(* Logix 5000 project; controller UOWHF_Vary Emulate 5570 rev 30.12; software revision 30.00; part 2 of 13 *)
(* tags used below, declared in another part *)
   UOWHF_Add_c : DINT;
   UOWHF_Msg : DINT[16];
   UOWHF_OutputMaxInd : DINT;
   UOWHF_Result : DINT[17];
(* MainProgram, continued *)

   		UOWHF_Result[2]:=UOWHF_Result[2] + 2135853958+UOWHF_Add_c;
   		UOWHF_Add_c.2:=UOWHF_Result[2].31;
   		UOWHF_Result[2].31:=0;
   		UOWHF_Result[3]:=UOWHF_Result[3] + 1732375759+UOWHF_Add_c;
   		UOWHF_Add_c.3:=UOWHF_Result[3].31;
   		UOWHF_Result[3].31:=0;
   		UOWHF_Result[4]:=UOWHF_Result[4] + 115158473+UOWHF_Add_c;
   		UOWHF_Add_c.4:=UOWHF_Result[4].31;
   		UOWHF_Result[4].31:=0;
   	End_If;
   	If UOWHF_Msg[4].[8] Then
   		UOWHF_Result[0]:=UOWHF_Result[0] + 1989798588+UOWHF_Add_c;
   		UOWHF_Add_c.0:=UOWHF_Result[0].31;
   		UOWHF_Result[0].31:=0;
   		UOWHF_Result[1]:=UOWHF_Result[1] + 591703516+UOWHF_Add_c;
   		UOWHF_Add_c.1:=UOWHF_Result[1].31;
   		UOWHF_Result[1].31:=0;
   		UOWHF_Result[2]:=UOWHF_Result[2] + 1328366246+UOWHF_Add_c;
   		UOWHF_Add_c.2:=UOWHF_Result[2].31;
   		UOWHF_Result[2].31:=0;
   		UOWHF_Result[3]:=UOWHF_Result[3] + 1055479196+UOWHF_Add_c;
   		UOWHF_Add_c.3:=UOWHF_Result[3].31;
   		UOWHF_Result[3].31:=0;
   		UOWHF_Result[4]:=UOWHF_Result[4] + 1638831242+UOWHF_Add_c;
   		UOWHF_Add_c.4:=UOWHF_Result[4].31;
   		UOWHF_Result[4].31:=0;
   	End_If;
   	If UOWHF_Msg[4].[9] Then
   		UOWHF_Result[0]:=UOWHF_Result[0] + 622406376+UOWHF_Add_c;
   		UOWHF_Add_c.0:=UOWHF_Result[0].31;
   		UOWHF_Result[0].31:=0;
   		UOWHF_Result[1]:=UOWHF_Result[1] + 302456745+UOWHF_Add_c;
   		UOWHF_Add_c.1:=UOWHF_Result[1].31;
   		UOWHF_Result[1].31:=0;
   		UOWHF_Result[2]:=UOWHF_Result[2] + 1004502914+UOWHF_Add_c;
   		UOWHF_Add_c.2:=UOWHF_Result[2].31;
   		UOWHF_Result[2].31:=0;
   		UOWHF_Result[3]:=UOWHF_Result[3] + 1944958998+UOWHF_Add_c;
   		UOWHF_Add_c.3:=UOWHF_Result[3].31;
   		UOWHF_Result[3].31:=0;
   		UOWHF_Result[4]:=UOWHF_Result[4] + 1457990763+UOWHF_Add_c;
   		UOWHF_Add_c.4:=UOWHF_Result[4].31;
   		UOWHF_Result[4].31:=0;
   	End_If;
   	If UOWHF_Msg[4].[10] Then
   		UOWHF_Result[0]:=UOWHF_Result[0] + 1190952435+UOWHF_Add_c;
   		UOWHF_Add_c.0:=UOWHF_Result[0].31;
   		UOWHF_Result[0].31:=0;
   		UOWHF_Result[1]:=UOWHF_Result[1] + 906321176+UOWHF_Add_c;
   		UOWHF_Add_c.1:=UOWHF_Result[1].31;
   		UOWHF_Result[1].31:=0;
   		UOWHF_Result[2]:=UOWHF_Result[2] + 1114856499+UOWHF_Add_c;
   		UOWHF_Add_c.2:=UOWHF_Result[2].31;
   		UOWHF_Result[2].31:=0;
   		UOWHF_Result[3]:=UOWHF_Result[3] + 2109990137+UOWHF_Add_c;
   		UOWHF_Add_c.3:=UOWHF_Result[3].31;
   		UOWHF_Result[3].31:=0;
   		UOWHF_Result[4]:=UOWHF_Result[4] + 2127466898+UOWHF_Add_c;
   		UOWHF_Add_c.4:=UOWHF_Result[4].31;
   		UOWHF_Result[4].31:=0;
   	End_If;
   	If UOWHF_Msg[4].[11] Then
   		UOWHF_Result[0]:=UOWHF_Result[0] + 1094778735+UOWHF_Add_c;
   		UOWHF_Add_c.0:=UOWHF_Result[0].31;
   		UOWHF_Result[0].31:=0;
   		UOWHF_Result[1]:=UOWHF_Result[1] + 920886974+UOWHF_Add_c;
   		UOWHF_Add_c.1:=UOWHF_Result[1].31;
   		UOWHF_Result[1].31:=0;
   		UOWHF_Result[2]:=UOWHF_Result[2] + 1275226437+UOWHF_Add_c;
   		UOWHF_Add_c.2:=UOWHF_Result[2].31;
   		UOWHF_Result[2].31:=0;
   		UOWHF_Result[3]:=UOWHF_Result[3] + 82556508+UOWHF_Add_c;
   		UOWHF_Add_c.3:=UOWHF_Result[3].31;
   		UOWHF_Result[3].31:=0;
   		UOWHF_Result[4]:=UOWHF_Result[4] + 977078858+UOWHF_Add_c;
   		UOWHF_Add_c.4:=UOWHF_Result[4].31;
   		UOWHF_Result[4].31:=0;
   	End_If;
   	If UOWHF_Msg[4].[12] Then
   		UOWHF_Result[0]:=UOWHF_Result[0] + 593744688+UOWHF_Add_c;
   		UOWHF_Add_c.0:=UOWHF_Result[0].31;
   		UOWHF_Result[0].31:=0;
   		UOWHF_Result[1]:=UOWHF_Result[1] + 1169255414+UOWHF_Add_c;
   		UOWHF_Add_c.1:=UOWHF_Result[1].31;
   		UOWHF_Result[1].31:=0;
   		UOWHF_Result[2]:=UOWHF_Result[2] + 51716405+UOWHF_Add_c;
   		UOWHF_Add_c.2:=UOWHF_Result[2].31;
   		UOWHF_Result[2].31:=0;
   		UOWHF_Result[3]:=UOWHF_Result[3] + 1207915051+UOWHF_Add_c;
   		UOWHF_Add_c.3:=UOWHF_Result[3].31;
   		UOWHF_Result[3].31:=0;
   		UOWHF_Result[4]:=UOWHF_Result[4] + 1842853883+UOWHF_Add_c;
   		UOWHF_Add_c.4:=UOWHF_Result[4].31;
   		UOWHF_Result[4].31:=0;
   	End_If;
   	If UOWHF_Msg[4].[13] Then
   		UOWHF_Result[0]:=UOWHF_Result[0] + 960750534+UOWHF_Add_c;
   		UOWHF_Add_c.0:=UOWHF_Result[0].31;
   		UOWHF_Result[0].31:=0;
   		UOWHF_Result[1]:=UOWHF_Result[1] + 581533276+UOWHF_Add_c;
   		UOWHF_Add_c.1:=UOWHF_Result[1].31;
   		UOWHF_Result[1].31:=0;
   		UOWHF_Result[2]:=UOWHF_Result[2] + 1726936368+UOWHF_Add_c;
   		UOWHF_Add_c.2:=UOWHF_Result[2].31;
   		UOWHF_Result[2].31:=0;
   		UOWHF_Result[3]:=UOWHF_Result[3] + 586011360+UOWHF_Add_c;
   		UOWHF_Add_c.3:=UOWHF_Result[3].31;
   		UOWHF_Result[3].31:=0;
   		UOWHF_Result[4]:=UOWHF_Result[4] + 1019866461+UOWHF_Add_c;
   		UOWHF_Add_c.4:=UOWHF_Result[4].31;
   		UOWHF_Result[4].31:=0;
   	End_If;
   	If UOWHF_Msg[4].[14] Then
   		UOWHF_Result[0]:=UOWHF_Result[0] + 867248205+UOWHF_Add_c;
   		UOWHF_Add_c.0:=UOWHF_Result[0].31;
   		UOWHF_Result[0].31:=0;
   		UOWHF_Result[1]:=UOWHF_Result[1] + 1887402509+UOWHF_Add_c;
   		UOWHF_Add_c.1:=UOWHF_Result[1].31;
   		UOWHF_Result[1].31:=0;
   		UOWHF_Result[2]:=UOWHF_Result[2] + 1521296444+UOWHF_Add_c;
   		UOWHF_Add_c.2:=UOWHF_Result[2].31;
   		UOWHF_Result[2].31:=0;
   		UOWHF_Result[3]:=UOWHF_Result[3] + 779741606+UOWHF_Add_c;
   		UOWHF_Add_c.3:=UOWHF_Result[3].31;
   		UOWHF_Result[3].31:=0;
   		UOWHF_Result[4]:=UOWHF_Result[4] + 1611229464+UOWHF_Add_c;
   		UOWHF_Add_c.4:=UOWHF_Result[4].31;
   		UOWHF_Result[4].31:=0;
   	End_If;
   	If UOWHF_Msg[4].[15] Then
   		UOWHF_Result[0]:=UOWHF_Result[0] + 1329140317+UOWHF_Add_c;
   		UOWHF_Add_c.0:=UOWHF_Result[0].31;
   		UOWHF_Result[0].31:=0;
   		UOWHF_Result[1]:=UOWHF_Result[1] + 1238656489+UOWHF_Add_c;
   		UOWHF_Add_c.1:=UOWHF_Result[1].31;
   		UOWHF_Result[1].31:=0;
   		UOWHF_Result[2]:=UOWHF_Result[2] + 252292269+UOWHF_Add_c;
   		UOWHF_Add_c.2:=UOWHF_Result[2].31;
   		UOWHF_Result[2].31:=0;
   		UOWHF_Result[3]:=UOWHF_Result[3] + 326259303+UOWHF_Add_c;
   		UOWHF_Add_c.3:=UOWHF_Result[3].31;
   		UOWHF_Result[3].31:=0;
   		UOWHF_Result[4]:=UOWHF_Result[4] + 469873786+UOWHF_Add_c;
   		UOWHF_Add_c.4:=UOWHF_Result[4].31;
   		UOWHF_Result[4].31:=0;
   	End_If;
   	If UOWHF_Msg[4].[16] Then
   		UOWHF_Result[0]:=UOWHF_Result[0] + 2017748157+UOWHF_Add_c;
   		UOWHF_Add_c.0:=UOWHF_Result[0].31;
   		UOWHF_Result[0].31:=0;
   		UOWHF_Result[1]:=UOWHF_Result[1] + 19496840+UOWHF_Add_c;
   		UOWHF_Add_c.1:=UOWHF_Result[1].31;
   		UOWHF_Result[1].31:=0;
   		UOWHF_Result[2]:=UOWHF_Result[2] + 1807187175+UOWHF_Add_c;
   		UOWHF_Add_c.2:=UOWHF_Result[2].31;
   		UOWHF_Result[2].31:=0;
   		UOWHF_Result[3]:=UOWHF_Result[3] + 293835404+UOWHF_Add_c;
   		UOWHF_Add_c.3:=UOWHF_Result[3].31;
   		UOWHF_Result[3].31:=0;
   		UOWHF_Result[4]:=UOWHF_Result[4] + 1565795281+UOWHF_Add_c;
   		UOWHF_Add_c.4:=UOWHF_Result[4].31;
   		UOWHF_Result[4].31:=0;
   	End_If;
   	If UOWHF_Msg[4].[17] Then
   		UOWHF_Result[0]:=UOWHF_Result[0] + 644949277+UOWHF_Add_c;
   		UOWHF_Add_c.0:=UOWHF_Result[0].31;
   		UOWHF_Result[0].31:=0;
   		UOWHF_Result[1]:=UOWHF_Result[1] + 917412774+UOWHF_Add_c;
   		UOWHF_Add_c.1:=UOWHF_Result[1].31;
   		UOWHF_Result[1].31:=0;
   		UOWHF_Result[2]:=UOWHF_Result[2] + 74925122+UOWHF_Add_c;
   		UOWHF_Add_c.2:=UOWHF_Result[2].31;
   		UOWHF_Result[2].31:=0;
   		UOWHF_Result[3]:=UOWHF_Result[3] + 406083723+UOWHF_Add_c;
   		UOWHF_Add_c.3:=UOWHF_Result[3].31;
   		UOWHF_Result[3].31:=0;
   		UOWHF_Result[4]:=UOWHF_Result[4] + 445412503+UOWHF_Add_c;
   		UOWHF_Add_c.4:=UOWHF_Result[4].31;
   		UOWHF_Result[4].31:=0;
   	End_If;
   	If UOWHF_Msg[4].[18] Then
   		UOWHF_Result[0]:=UOWHF_Result[0] + 469282993+UOWHF_Add_c;
   		UOWHF_Add_c.0:=UOWHF_Result[0].31;
   		UOWHF_Result[0].31:=0;
   		UOWHF_Result[1]:=UOWHF_Result[1] + 429116135+UOWHF_Add_c;
   		UOWHF_Add_c.1:=UOWHF_Result[1].31;
   		UOWHF_Result[1].31:=0;
   		UOWHF_Result[2]:=UOWHF_Result[2] + 2025571244+UOWHF_Add_c;
   		UOWHF_Add_c.2:=UOWHF_Result[2].31;
   		UOWHF_Result[2].31:=0;
   		UOWHF_Result[3]:=UOWHF_Result[3] + 1523762277+UOWHF_Add_c;
   		UOWHF_Add_c.3:=UOWHF_Result[3].31;
   		UOWHF_Result[3].31:=0;
   		UOWHF_Result[4]:=UOWHF_Result[4] + 1908737666+UOWHF_Add_c;
   		UOWHF_Add_c.4:=UOWHF_Result[4].31;
   		UOWHF_Result[4].31:=0;
   	End_If;
   	If UOWHF_Msg[4].[19] Then
   		UOWHF_Result[0]:=UOWHF_Result[0] + 1510848022+UOWHF_Add_c;
   		UOWHF_Add_c.0:=UOWHF_Result[0].31;
   		UOWHF_Result[0].31:=0;
   		UOWHF_Result[1]:=UOWHF_Result[1] + 256825122+UOWHF_Add_c;
   		UOWHF_Add_c.1:=UOWHF_Result[1].31;
   		UOWHF_Result[1].31:=0;
   		UOWHF_Result[2]:=UOWHF_Result[2] + 1516475094+UOWHF_Add_c;
   		UOWHF_Add_c.2:=UOWHF_Result[2].31;
   		UOWHF_Result[2].31:=0;
   		UOWHF_Result[3]:=UOWHF_Result[3] + 1288161802+UOWHF_Add_c;
   		UOWHF_Add_c.3:=UOWHF_Result[3].31;
   		UOWHF_Result[3].31:=0;
   		UOWHF_Result[4]:=UOWHF_Result[4] + 366249542+UOWHF_Add_c;
   		UOWHF_Add_c.4:=UOWHF_Result[4].31;
   		UOWHF_Result[4].31:=0;
   	End_If;
   	If UOWHF_Msg[4].[20] Then
   		UOWHF_Result[0]:=UOWHF_Result[0] + 1574992729+UOWHF_Add_c;
   		UOWHF_Add_c.0:=UOWHF_Result[0].31;
   		UOWHF_Result[0].31:=0;
   		UOWHF_Result[1]:=UOWHF_Result[1] + 274898417+UOWHF_Add_c;
   		UOWHF_Add_c.1:=UOWHF_Result[1].31;
   		UOWHF_Result[1].31:=0;
   		UOWHF_Result[2]:=UOWHF_Result[2] + 1217972673+UOWHF_Add_c;
   		UOWHF_Add_c.2:=UOWHF_Result[2].31;
   		UOWHF_Result[2].31:=0;
   		UOWHF_Result[3]:=UOWHF_Result[3] + 491443084+UOWHF_Add_c;
   		UOWHF_Add_c.3:=UOWHF_Result[3].31;
   		UOWHF_Result[3].31:=0;
   		UOWHF_Result[4]:=UOWHF_Result[4] + 1677131526+UOWHF_Add_c;
   		UOWHF_Add_c.4:=UOWHF_Result[4].31;
   		UOWHF_Result[4].31:=0;
   	End_If;
   	If UOWHF_Msg[4].[21] Then
   		UOWHF_Result[0]:=UOWHF_Result[0] + 1458801108+UOWHF_Add_c;
   		UOWHF_Add_c.0:=UOWHF_Result[0].31;
   		UOWHF_Result[0].31:=0;
   		UOWHF_Result[1]:=UOWHF_Result[1] + 1008833420+UOWHF_Add_c;
   		UOWHF_Add_c.1:=UOWHF_Result[1].31;
   		UOWHF_Result[1].31:=0;
   		UOWHF_Result[2]:=UOWHF_Result[2] + 6669131+UOWHF_Add_c;
   		UOWHF_Add_c.2:=UOWHF_Result[2].31;
   		UOWHF_Result[2].31:=0;
   		UOWHF_Result[3]:=UOWHF_Result[3] + 606622791+UOWHF_Add_c;
   		UOWHF_Add_c.3:=UOWHF_Result[3].31;
   		UOWHF_Result[3].31:=0;
   		UOWHF_Result[4]:=UOWHF_Result[4] + 1662810500+UOWHF_Add_c;
   		UOWHF_Add_c.4:=UOWHF_Result[4].31;
   		UOWHF_Result[4].31:=0;
   	End_If;
   	If UOWHF_Msg[4].[22] Then
   		UOWHF_Result[0]:=UOWHF_Result[0] + 929898449+UOWHF_Add_c;
   		UOWHF_Add_c.0:=UOWHF_Result[0].31;
   		UOWHF_Result[0].31:=0;
   		UOWHF_Result[1]:=UOWHF_Result[1] + 1134852805+UOWHF_Add_c;
   		UOWHF_Add_c.1:=UOWHF_Result[1].31;
   		UOWHF_Result[1].31:=0;
   		UOWHF_Result[2]:=UOWHF_Result[2] + 1313816737+UOWHF_Add_c;
   		UOWHF_Add_c.2:=UOWHF_Result[2].31;
   		UOWHF_Result[2].31:=0;
   		UOWHF_Result[3]:=UOWHF_Result[3] + 1450371462+UOWHF_Add_c;
   		UOWHF_Add_c.3:=UOWHF_Result[3].31;
   		UOWHF_Result[3].31:=0;
   		UOWHF_Result[4]:=UOWHF_Result[4] + 1409338575+UOWHF_Add_c;
   		UOWHF_Add_c.4:=UOWHF_Result[4].31;
   		UOWHF_Result[4].31:=0;
   	End_If;
   	If UOWHF_Msg[4].[23] Then
   		UOWHF_Result[0]:=UOWHF_Result[0] + 1696773702+UOWHF_Add_c;
   		UOWHF_Add_c.0:=UOWHF_Result[0].31;
   		UOWHF_Result[0].31:=0;
   		UOWHF_Result[1]:=UOWHF_Result[1] + 1574239672+UOWHF_Add_c;
   		UOWHF_Add_c.1:=UOWHF_Result[1].31;
   		UOWHF_Result[1].31:=0;
   		UOWHF_Result[2]:=UOWHF_Result[2] + 845690239+UOWHF_Add_c;
   		UOWHF_Add_c.2:=UOWHF_Result[2].31;
   		UOWHF_Result[2].31:=0;
   		UOWHF_Result[3]:=UOWHF_Result[3] + 301138788+UOWHF_Add_c;
   		UOWHF_Add_c.3:=UOWHF_Result[3].31;
   		UOWHF_Result[3].31:=0;
   		UOWHF_Result[4]:=UOWHF_Result[4] + 953256044+UOWHF_Add_c;
   		UOWHF_Add_c.4:=UOWHF_Result[4].31;
   		UOWHF_Result[4].31:=0;
   	End_If;
   	If UOWHF_Msg[4].[24] Then
   		UOWHF_Result[0]:=UOWHF_Result[0] + 51899107+UOWHF_Add_c;
   		UOWHF_Add_c.0:=UOWHF_Result[0].31;
   		UOWHF_Result[0].31:=0;
   		UOWHF_Result[1]:=UOWHF_Result[1] + 286317975+UOWHF_Add_c;
   		UOWHF_Add_c.1:=UOWHF_Result[1].31;
   		UOWHF_Result[1].31:=0;
   		UOWHF_Result[2]:=UOWHF_Result[2] + 841734893+UOWHF_Add_c;
   		UOWHF_Add_c.2:=UOWHF_Result[2].31;
   		UOWHF_Result[2].31:=0;
   		UOWHF_Result[3]:=UOWHF_Result[3] + 902319505+UOWHF_Add_c;
   		UOWHF_Add_c.3:=UOWHF_Result[3].31;
   		UOWHF_Result[3].31:=0;
   		UOWHF_Result[4]:=UOWHF_Result[4] + 1996737543+UOWHF_Add_c;
   		UOWHF_Add_c.4:=UOWHF_Result[4].31;
   		UOWHF_Result[4].31:=0;
   	End_If;
   	If UOWHF_Msg[4].[25] Then
   		UOWHF_Result[0]:=UOWHF_Result[0] + 299129534+UOWHF_Add_c;
   		UOWHF_Add_c.0:=UOWHF_Result[0].31;
   		UOWHF_Result[0].31:=0;
   		UOWHF_Result[1]:=UOWHF_Result[1] + 1540449511+UOWHF_Add_c;
   		UOWHF_Add_c.1:=UOWHF_Result[1].31;
   		UOWHF_Result[1].31:=0;
   		UOWHF_Result[2]:=UOWHF_Result[2] + 323357098+UOWHF_Add_c;
   		UOWHF_Add_c.2:=UOWHF_Result[2].31;
   		UOWHF_Result[2].31:=0;
   		UOWHF_Result[3]:=UOWHF_Result[3] + 605016071+UOWHF_Add_c;
   		UOWHF_Add_c.3:=UOWHF_Result[3].31;
   		UOWHF_Result[3].31:=0;
   		UOWHF_Result[4]:=UOWHF_Result[4] + 627496508+UOWHF_Add_c;
   		UOWHF_Add_c.4:=UOWHF_Result[4].31;
   		UOWHF_Result[4].31:=0;
   	End_If;
   	If UOWHF_Msg[4].[26] Then
   		UOWHF_Result[0]:=UOWHF_Result[0] + 930496525+UOWHF_Add_c;
   		UOWHF_Add_c.0:=UOWHF_Result[0].31;
   		UOWHF_Result[0].31:=0;
   		UOWHF_Result[1]:=UOWHF_Result[1] + 242034892+UOWHF_Add_c;
   		UOWHF_Add_c.1:=UOWHF_Result[1].31;
   		UOWHF_Result[1].31:=0;
   		UOWHF_Result[2]:=UOWHF_Result[2] + 613467940+UOWHF_Add_c;
   		UOWHF_Add_c.2:=UOWHF_Result[2].31;
   		UOWHF_Result[2].31:=0;
   		UOWHF_Result[3]:=UOWHF_Result[3] + 385508360+UOWHF_Add_c;
   		UOWHF_Add_c.3:=UOWHF_Result[3].31;
   		UOWHF_Result[3].31:=0;
   		UOWHF_Result[4]:=UOWHF_Result[4] + 1770337894+UOWHF_Add_c;
   		UOWHF_Add_c.4:=UOWHF_Result[4].31;
   		UOWHF_Result[4].31:=0;
   	End_If;
   	If UOWHF_Msg[4].[27] Then
   		UOWHF_Result[0]:=UOWHF_Result[0] + 2063144581+UOWHF_Add_c;
   		UOWHF_Add_c.0:=UOWHF_Result[0].31;
   		UOWHF_Result[0].31:=0;
   		UOWHF_Result[1]:=UOWHF_Result[1] + 1679769568+UOWHF_Add_c;
   		UOWHF_Add_c.1:=UOWHF_Result[1].31;
   		UOWHF_Result[1].31:=0;
   		UOWHF_Result[2]:=UOWHF_Result[2] + 2137628573+UOWHF_Add_c;
   		UOWHF_Add_c.2:=UOWHF_Result[2].31;
   		UOWHF_Result[2].31:=0;
   		UOWHF_Result[3]:=UOWHF_Result[3] + 778926313+UOWHF_Add_c;
   		UOWHF_Add_c.3:=UOWHF_Result[3].31;
   		UOWHF_Result[3].31:=0;
   		UOWHF_Result[4]:=UOWHF_Result[4] + 1705142262+UOWHF_Add_c;
   		UOWHF_Add_c.4:=UOWHF_Result[4].31;
   		UOWHF_Result[4].31:=0;
   	End_If;
   	If UOWHF_Msg[4].[28] Then
   		UOWHF_Result[0]:=UOWHF_Result[0] + 223464317+UOWHF_Add_c;
   		UOWHF_Add_c.0:=UOWHF_Result[0].31;
   		UOWHF_Result[0].31:=0;
   		UOWHF_Result[1]:=UOWHF_Result[1] + 154890765+UOWHF_Add_c;
   		UOWHF_Add_c.1:=UOWHF_Result[1].31;
   		UOWHF_Result[1].31:=0;
   		UOWHF_Result[2]:=UOWHF_Result[2] + 866520135+UOWHF_Add_c;
   		UOWHF_Add_c.2:=UOWHF_Result[2].31;
   		UOWHF_Result[2].31:=0;
   		UOWHF_Result[3]:=UOWHF_Result[3] + 1732824316+UOWHF_Add_c;
   		UOWHF_Add_c.3:=UOWHF_Result[3].31;
   		UOWHF_Result[3].31:=0;
   		UOWHF_Result[4]:=UOWHF_Result[4] + 622807513+UOWHF_Add_c;
   		UOWHF_Add_c.4:=UOWHF_Result[4].31;
   		UOWHF_Result[4].31:=0;
   	End_If;
   	If UOWHF_Msg[4].[29] Then
   		UOWHF_Result[0]:=UOWHF_Result[0] + 469565239+UOWHF_Add_c;
   		UOWHF_Add_c.0:=UOWHF_Result[0].31;
   		UOWHF_Result[0].31:=0;
   		UOWHF_Result[1]:=UOWHF_Result[1] + 1133898399+UOWHF_Add_c;
   		UOWHF_Add_c.1:=UOWHF_Result[1].31;
   		UOWHF_Result[1].31:=0;
   		UOWHF_Result[2]:=UOWHF_Result[2] + 2080362872+UOWHF_Add_c;
   		UOWHF_Add_c.2:=UOWHF_Result[2].31;
   		UOWHF_Result[2].31:=0;
   		UOWHF_Result[3]:=UOWHF_Result[3] + 1351452134+UOWHF_Add_c;
   		UOWHF_Add_c.3:=UOWHF_Result[3].31;
   		UOWHF_Result[3].31:=0;
   		UOWHF_Result[4]:=UOWHF_Result[4] + 1256652494+UOWHF_Add_c;
   		UOWHF_Add_c.4:=UOWHF_Result[4].31;
   		UOWHF_Result[4].31:=0;
   	End_If;
   	If UOWHF_Msg[4].[30] Then
   		UOWHF_Result[0]:=UOWHF_Result[0] + 139067637+UOWHF_Add_c;
   		UOWHF_Add_c.0:=UOWHF_Result[0].31;
   		UOWHF_Result[0].31:=0;
   		UOWHF_Result[1]:=UOWHF_Result[1] + 130304763+UOWHF_Add_c;
   		UOWHF_Add_c.1:=UOWHF_Result[1].31;
   		UOWHF_Result[1].31:=0;
   		UOWHF_Result[2]:=UOWHF_Result[2] + 1233288998+UOWHF_Add_c;
   		UOWHF_Add_c.2:=UOWHF_Result[2].31;
   		UOWHF_Result[2].31:=0;
   		UOWHF_Result[3]:=UOWHF_Result[3] + 314279374+UOWHF_Add_c;
   		UOWHF_Add_c.3:=UOWHF_Result[3].31;
   		UOWHF_Result[3].31:=0;
   		UOWHF_Result[4]:=UOWHF_Result[4] + 1142265410+UOWHF_Add_c;
   		UOWHF_Add_c.4:=UOWHF_Result[4].31;
   		UOWHF_Result[4].31:=0;
   	End_If;
   	If UOWHF_Msg[4].[31] Then
   		UOWHF_Result[0]:=UOWHF_Result[0] + 600121605+UOWHF_Add_c;
   		UOWHF_Add_c.0:=UOWHF_Result[0].31;
   		UOWHF_Result[0].31:=0;
   		UOWHF_Result[1]:=UOWHF_Result[1] + 1762194152+UOWHF_Add_c;
   		UOWHF_Add_c.1:=UOWHF_Result[1].31;
   		UOWHF_Result[1].31:=0;
   		UOWHF_Result[2]:=UOWHF_Result[2] + 1169274486+UOWHF_Add_c;
   		UOWHF_Add_c.2:=UOWHF_Result[2].31;
   		UOWHF_Result[2].31:=0;
   		UOWHF_Result[3]:=UOWHF_Result[3] + 2110531411+UOWHF_Add_c;
   		UOWHF_Add_c.3:=UOWHF_Result[3].31;
   		UOWHF_Result[3].31:=0;
   		UOWHF_Result[4]:=UOWHF_Result[4] + 863289396+UOWHF_Add_c;
   		UOWHF_Add_c.4:=UOWHF_Result[4].31;
   		UOWHF_Result[4].31:=0;
   	End_If;
   	If UOWHF_Msg[5].[0] Then
   		UOWHF_Result[0]:=UOWHF_Result[0] + 1573571782+UOWHF_Add_c;
   		UOWHF_Add_c.0:=UOWHF_Result[0].31;
   		UOWHF_Result[0].31:=0;
   		UOWHF_Result[1]:=UOWHF_Result[1] + 1156496734+UOWHF_Add_c;
   		UOWHF_Add_c.1:=UOWHF_Result[1].31;
   		UOWHF_Result[1].31:=0;
   		UOWHF_Result[2]:=UOWHF_Result[2] + 1922217724+UOWHF_Add_c;
   		UOWHF_Add_c.2:=UOWHF_Result[2].31;
   		UOWHF_Result[2].31:=0;
   		UOWHF_Result[3]:=UOWHF_Result[3] + 1472440733+UOWHF_Add_c;
   		UOWHF_Add_c.3:=UOWHF_Result[3].31;
   		UOWHF_Result[3].31:=0;
   		UOWHF_Result[4]:=UOWHF_Result[4] + 1603570212+UOWHF_Add_c;
   		UOWHF_Add_c.4:=UOWHF_Result[4].31;
   		UOWHF_Result[4].31:=0;
   	End_If;
   	If UOWHF_Msg[5].[1] Then
   		UOWHF_Result[0]:=UOWHF_Result[0] + 1081646203+UOWHF_Add_c;
   		UOWHF_Add_c.0:=UOWHF_Result[0].31;
   		UOWHF_Result[0].31:=0;
   		UOWHF_Result[1]:=UOWHF_Result[1] + 897382485+UOWHF_Add_c;
   		UOWHF_Add_c.1:=UOWHF_Result[1].31;
   		UOWHF_Result[1].31:=0;
   		UOWHF_Result[2]:=UOWHF_Result[2] + 1891296415+UOWHF_Add_c;
   		UOWHF_Add_c.2:=UOWHF_Result[2].31;
   		UOWHF_Result[2].31:=0;
   		UOWHF_Result[3]:=UOWHF_Result[3] + 531871977+UOWHF_Add_c;
   		UOWHF_Add_c.3:=UOWHF_Result[3].31;
   		UOWHF_Result[3].31:=0;
   		UOWHF_Result[4]:=UOWHF_Result[4] + 1737698500+UOWHF_Add_c;
   		UOWHF_Add_c.4:=UOWHF_Result[4].31;
   		UOWHF_Result[4].31:=0;
   	End_If;
   	If UOWHF_Msg[5].[2] Then
   		UOWHF_Result[0]:=UOWHF_Result[0] + 188343515+UOWHF_Add_c;
   		UOWHF_Add_c.0:=UOWHF_Result[0].31;
   		UOWHF_Result[0].31:=0;
   		UOWHF_Result[1]:=UOWHF_Result[1] + 626004248+UOWHF_Add_c;
   		UOWHF_Add_c.1:=UOWHF_Result[1].31;
   		UOWHF_Result[1].31:=0;
   		UOWHF_Result[2]:=UOWHF_Result[2] + 1577949949+UOWHF_Add_c;
   		UOWHF_Add_c.2:=UOWHF_Result[2].31;
   		UOWHF_Result[2].31:=0;
   		UOWHF_Result[3]:=UOWHF_Result[3] + 1536216209+UOWHF_Add_c;
   		UOWHF_Add_c.3:=UOWHF_Result[3].31;
   		UOWHF_Result[3].31:=0;
   		UOWHF_Result[4]:=UOWHF_Result[4] + 1377657699+UOWHF_Add_c;
   		UOWHF_Add_c.4:=UOWHF_Result[4].31;
   		UOWHF_Result[4].31:=0;
   	End_If;
   	If UOWHF_Msg[5].[3] Then
   		UOWHF_Result[0]:=UOWHF_Result[0] + 1561195711+UOWHF_Add_c;
   		UOWHF_Add_c.0:=UOWHF_Result[0].31;
   		UOWHF_Result[0].31:=0;
   		UOWHF_Result[1]:=UOWHF_Result[1] + 223853766+UOWHF_Add_c;
   		UOWHF_Add_c.1:=UOWHF_Result[1].31;
   		UOWHF_Result[1].31:=0;
   		UOWHF_Result[2]:=UOWHF_Result[2] + 1814003587+UOWHF_Add_c;
   		UOWHF_Add_c.2:=UOWHF_Result[2].31;
   		UOWHF_Result[2].31:=0;
   		UOWHF_Result[3]:=UOWHF_Result[3] + 274097477+UOWHF_Add_c;
   		UOWHF_Add_c.3:=UOWHF_Result[3].31;
   		UOWHF_Result[3].31:=0;
   		UOWHF_Result[4]:=UOWHF_Result[4] + 1280958193+UOWHF_Add_c;
   		UOWHF_Add_c.4:=UOWHF_Result[4].31;
   		UOWHF_Result[4].31:=0;
   	End_If;
   	If UOWHF_Msg[5].[4] Then
   		UOWHF_Result[0]:=UOWHF_Result[0] + 532570630+UOWHF_Add_c;
   		UOWHF_Add_c.0:=UOWHF_Result[0].31;
   		UOWHF_Result[0].31:=0;
   		UOWHF_Result[1]:=UOWHF_Result[1] + 883659870+UOWHF_Add_c;
   		UOWHF_Add_c.1:=UOWHF_Result[1].31;
   		UOWHF_Result[1].31:=0;
   		UOWHF_Result[2]:=UOWHF_Result[2] + 479800569+UOWHF_Add_c;
   		UOWHF_Add_c.2:=UOWHF_Result[2].31;
   		UOWHF_Result[2].31:=0;
   		UOWHF_Result[3]:=UOWHF_Result[3] + 75520038+UOWHF_Add_c;
   		UOWHF_Add_c.3:=UOWHF_Result[3].31;
   		UOWHF_Result[3].31:=0;
   		UOWHF_Result[4]:=UOWHF_Result[4] + 117000370+UOWHF_Add_c;
   		UOWHF_Add_c.4:=UOWHF_Result[4].31;
   		UOWHF_Result[4].31:=0;
   	End_If;
   	If UOWHF_Msg[5].[5] Then
   		UOWHF_Result[0]:=UOWHF_Result[0] + 719275818+UOWHF_Add_c;
   		UOWHF_Add_c.0:=UOWHF_Result[0].31;
   		UOWHF_Result[0].31:=0;
   		UOWHF_Result[1]:=UOWHF_Result[1] + 878778090+UOWHF_Add_c;
   		UOWHF_Add_c.1:=UOWHF_Result[1].31;
   		UOWHF_Result[1].31:=0;
   		UOWHF_Result[2]:=UOWHF_Result[2] + 1579901234+UOWHF_Add_c;
   		UOWHF_Add_c.2:=UOWHF_Result[2].31;
   		UOWHF_Result[2].31:=0;
   		UOWHF_Result[3]:=UOWHF_Result[3] + 1303455866+UOWHF_Add_c;
   		UOWHF_Add_c.3:=UOWHF_Result[3].31;
   		UOWHF_Result[3].31:=0;
   		UOWHF_Result[4]:=UOWHF_Result[4] + 1769591178+UOWHF_Add_c;
   		UOWHF_Add_c.4:=UOWHF_Result[4].31;
   		UOWHF_Result[4].31:=0;
   	End_If;
   	If UOWHF_Msg[5].[6] Then
   		UOWHF_Result[0]:=UOWHF_Result[0] + 196695134+UOWHF_Add_c;
   		UOWHF_Add_c.0:=UOWHF_Result[0].31;
   		UOWHF_Result[0].31:=0;
   		UOWHF_Result[1]:=UOWHF_Result[1] + 1352456716+UOWHF_Add_c;
   		UOWHF_Add_c.1:=UOWHF_Result[1].31;
   		UOWHF_Result[1].31:=0;
   		UOWHF_Result[2]:=UOWHF_Result[2] + 496301287+UOWHF_Add_c;
   		UOWHF_Add_c.2:=UOWHF_Result[2].31;
   		UOWHF_Result[2].31:=0;
   		UOWHF_Result[3]:=UOWHF_Result[3] + 1532761137+UOWHF_Add_c;
   		UOWHF_Add_c.3:=UOWHF_Result[3].31;
   		UOWHF_Result[3].31:=0;
   		UOWHF_Result[4]:=UOWHF_Result[4] + 51579917+UOWHF_Add_c;
   		UOWHF_Add_c.4:=UOWHF_Result[4].31;
   		UOWHF_Result[4].31:=0;
   	End_If;
   	If UOWHF_Msg[5].[7] Then
   		UOWHF_Result[0]:=UOWHF_Result[0] + 1250982478+UOWHF_Add_c;
   		UOWHF_Add_c.0:=UOWHF_Result[0].31;
   		UOWHF_Result[0].31:=0;
   		UOWHF_Result[1]:=UOWHF_Result[1] + 2035409170+UOWHF_Add_c;
   		UOWHF_Add_c.1:=UOWHF_Result[1].31;
   		UOWHF_Result[1].31:=0;
   		UOWHF_Result[2]:=UOWHF_Result[2] + 1771335087+UOWHF_Add_c;
   		UOWHF_Add_c.2:=UOWHF_Result[2].31;
   		UOWHF_Result[2].31:=0;
   		UOWHF_Result[3]:=UOWHF_Result[3] + 546944966+UOWHF_Add_c;
   		UOWHF_Add_c.3:=UOWHF_Result[3].31;
   		UOWHF_Result[3].31:=0;
   		UOWHF_Result[4]:=UOWHF_Result[4] + 285453755+UOWHF_Add_c;
   		UOWHF_Add_c.4:=UOWHF_Result[4].31;
   		UOWHF_Result[4].31:=0;
   	End_If;
   	If UOWHF_Msg[5].[8] Then
   		UOWHF_Result[0]:=UOWHF_Result[0] + 1954924621+UOWHF_Add_c;
   		UOWHF_Add_c.0:=UOWHF_Result[0].31;
   		UOWHF_Result[0].31:=0;
   		UOWHF_Result[1]:=UOWHF_Result[1] + 1539545990+UOWHF_Add_c;
   		UOWHF_Add_c.1:=UOWHF_Result[1].31;
   		UOWHF_Result[1].31:=0;
   		UOWHF_Result[2]:=UOWHF_Result[2] + 19863553+UOWHF_Add_c;
   		UOWHF_Add_c.2:=UOWHF_Result[2].31;
   		UOWHF_Result[2].31:=0;
   		UOWHF_Result[3]:=UOWHF_Result[3] + 2001043044+UOWHF_Add_c;
   		UOWHF_Add_c.3:=UOWHF_Result[3].31;
   		UOWHF_Result[3].31:=0;
   		UOWHF_Result[4]:=UOWHF_Result[4] + 506173703+UOWHF_Add_c;
   		UOWHF_Add_c.4:=UOWHF_Result[4].31;
   		UOWHF_Result[4].31:=0;
   	End_If;
   	If UOWHF_Msg[5].[9] Then
   		UOWHF_Result[0]:=UOWHF_Result[0] + 726827605+UOWHF_Add_c;
   		UOWHF_Add_c.0:=UOWHF_Result[0].31;
   		UOWHF_Result[0].31:=0;
   		UOWHF_Result[1]:=UOWHF_Result[1] + 345457676+UOWHF_Add_c;
   		UOWHF_Add_c.1:=UOWHF_Result[1].31;
   		UOWHF_Result[1].31:=0;
   		UOWHF_Result[2]:=UOWHF_Result[2] + 1181066952+UOWHF_Add_c;
   		UOWHF_Add_c.2:=UOWHF_Result[2].31;
   		UOWHF_Result[2].31:=0;
   		UOWHF_Result[3]:=UOWHF_Result[3] + 399489837+UOWHF_Add_c;
   		UOWHF_Add_c.3:=UOWHF_Result[3].31;
   		UOWHF_Result[3].31:=0;
   		UOWHF_Result[4]:=UOWHF_Result[4] + 345723933+UOWHF_Add_c;
   		UOWHF_Add_c.4:=UOWHF_Result[4].31;
   		UOWHF_Result[4].31:=0;
   	End_If;
   	If UOWHF_Msg[5].[10] Then
   		UOWHF_Result[0]:=UOWHF_Result[0] + 376333595+UOWHF_Add_c;
   		UOWHF_Add_c.0:=UOWHF_Result[0].31;
   		UOWHF_Result[0].31:=0;
   		UOWHF_Result[1]:=UOWHF_Result[1] + 655993442+UOWHF_Add_c;
   		UOWHF_Add_c.1:=UOWHF_Result[1].31;
   		UOWHF_Result[1].31:=0;
   		UOWHF_Result[2]:=UOWHF_Result[2] + 1300987572+UOWHF_Add_c;
   		UOWHF_Add_c.2:=UOWHF_Result[2].31;
   		UOWHF_Result[2].31:=0;
   		UOWHF_Result[3]:=UOWHF_Result[3] + 744685865+UOWHF_Add_c;
   		UOWHF_Add_c.3:=UOWHF_Result[3].31;
   		UOWHF_Result[3].31:=0;
   		UOWHF_Result[4]:=UOWHF_Result[4] + 1482881180+UOWHF_Add_c;
   		UOWHF_Add_c.4:=UOWHF_Result[4].31;
   		UOWHF_Result[4].31:=0;
   	End_If;
   	If UOWHF_Msg[5].[11] Then
   		UOWHF_Result[0]:=UOWHF_Result[0] + 136189820+UOWHF_Add_c;
   		UOWHF_Add_c.0:=UOWHF_Result[0].31;
   		UOWHF_Result[0].31:=0;
   		UOWHF_Result[1]:=UOWHF_Result[1] + 1112761140+UOWHF_Add_c;
   		UOWHF_Add_c.1:=UOWHF_Result[1].31;
   		UOWHF_Result[1].31:=0;
   		UOWHF_Result[2]:=UOWHF_Result[2] + 1915046367+UOWHF_Add_c;
   		UOWHF_Add_c.2:=UOWHF_Result[2].31;
   		UOWHF_Result[2].31:=0;
   		UOWHF_Result[3]:=UOWHF_Result[3] + 1660983898+UOWHF_Add_c;
   		UOWHF_Add_c.3:=UOWHF_Result[3].31;
   		UOWHF_Result[3].31:=0;
   		UOWHF_Result[4]:=UOWHF_Result[4] + 1697634729+UOWHF_Add_c;
   		UOWHF_Add_c.4:=UOWHF_Result[4].31;
   		UOWHF_Result[4].31:=0;
   	End_If;
   	If UOWHF_Msg[5].[12] Then
   		UOWHF_Result[0]:=UOWHF_Result[0] + 556388719+UOWHF_Add_c;
   		UOWHF_Add_c.0:=UOWHF_Result[0].31;
   		UOWHF_Result[0].31:=0;
   		UOWHF_Result[1]:=UOWHF_Result[1] + 1862688541+UOWHF_Add_c;
   		UOWHF_Add_c.1:=UOWHF_Result[1].31;
   		UOWHF_Result[1].31:=0;
   		UOWHF_Result[2]:=UOWHF_Result[2] + 484621113+UOWHF_Add_c;
   		UOWHF_Add_c.2:=UOWHF_Result[2].31;
   		UOWHF_Result[2].31:=0;
   		UOWHF_Result[3]:=UOWHF_Result[3] + 393036979+UOWHF_Add_c;
   		UOWHF_Add_c.3:=UOWHF_Result[3].31;
   		UOWHF_Result[3].31:=0;
   		UOWHF_Result[4]:=UOWHF_Result[4] + 1415012869+UOWHF_Add_c;
   		UOWHF_Add_c.4:=UOWHF_Result[4].31;
   		UOWHF_Result[4].31:=0;
   	End_If;
   	If UOWHF_Msg[5].[13] Then
   		UOWHF_Result[0]:=UOWHF_Result[0] + 1972057419+UOWHF_Add_c;
   		UOWHF_Add_c.0:=UOWHF_Result[0].31;
   		UOWHF_Result[0].31:=0;
   		UOWHF_Result[1]:=UOWHF_Result[1] + 1673453536+UOWHF_Add_c;
   		UOWHF_Add_c.1:=UOWHF_Result[1].31;
   		UOWHF_Result[1].31:=0;
   		UOWHF_Result[2]:=UOWHF_Result[2] + 1268609640+UOWHF_Add_c;
   		UOWHF_Add_c.2:=UOWHF_Result[2].31;
   		UOWHF_Result[2].31:=0;
   		UOWHF_Result[3]:=UOWHF_Result[3] + 972799653+UOWHF_Add_c;
   		UOWHF_Add_c.3:=UOWHF_Result[3].31;
   		UOWHF_Result[3].31:=0;
   		UOWHF_Result[4]:=UOWHF_Result[4] + 527216737+UOWHF_Add_c;
   		UOWHF_Add_c.4:=UOWHF_Result[4].31;
   		UOWHF_Result[4].31:=0;
   	End_If;
   	If UOWHF_Msg[5].[14] Then
   		UOWHF_Result[0]:=UOWHF_Result[0] + 1813383740+UOWHF_Add_c;
   		UOWHF_Add_c.0:=UOWHF_Result[0].31;
   		UOWHF_Result[0].31:=0;
   		UOWHF_Result[1]:=UOWHF_Result[1] + 2015396043+UOWHF_Add_c;
   		UOWHF_Add_c.1:=UOWHF_Result[1].31;
   		UOWHF_Result[1].31:=0;
   		UOWHF_Result[2]:=UOWHF_Result[2] + 1315693252+UOWHF_Add_c;
   		UOWHF_Add_c.2:=UOWHF_Result[2].31;
   		UOWHF_Result[2].31:=0;
   		UOWHF_Result[3]:=UOWHF_Result[3] + 1148760085+UOWHF_Add_c;
   		UOWHF_Add_c.3:=UOWHF_Result[3].31;
   		UOWHF_Result[3].31:=0;
   		UOWHF_Result[4]:=UOWHF_Result[4] + 1548609049+UOWHF_Add_c;
   		UOWHF_Add_c.4:=UOWHF_Result[4].31;
   		UOWHF_Result[4].31:=0;
   	End_If;
   	If UOWHF_Msg[5].[15] Then
   		UOWHF_Result[0]:=UOWHF_Result[0] + 1194474809+UOWHF_Add_c;
   		UOWHF_Add_c.0:=UOWHF_Result[0].31;
   		UOWHF_Result[0].31:=0;
   		UOWHF_Result[1]:=UOWHF_Result[1] + 808421095+UOWHF_Add_c;
   		UOWHF_Add_c.1:=UOWHF_Result[1].31;
   		UOWHF_Result[1].31:=0;